   3396: 'Carrier 53 CB02122 Tripped', class No Acknowledgement, trigger "DB302_HMI_Faults_Carrier53_Faults_0" bit 3
   3397: 'Carrier 53 CB02123 Tripped', class No Acknowledgement, trigger "DB302_HMI_Faults_Carrier53_Faults_0" bit 4
   3398: 'Carrier 53 AUX1 CB Tripped', class No Acknowledgement, trigger "DB302_HMI_Faults_Carrier53_Faults_0" bit 5
   3399: 'Carrier 53 AUX2 CB Tripped', class No Acknowledgement, trigger "DB302_HMI_Faults_Carrier53_Faults_0" bit 6
   3400: 'Carrier 53 PLC Not Communicating', class No Acknowledgement, trigger "DB302_HMI_Faults_Carrier53_Faults_0" bit 7
   3401: 'Carrier 53 Safe Input Card Fault', class No Acknowledgement, trigger "DB302_HMI_Faults_Carrier53_Faults_0" bit 8
   3402: 'Carrier 53 Safe Output Card Fault', class No Acknowledgement, trigger "DB302_HMI_Faults_Carrier53_Faults_0" bit 9
   3403: 'Carrier 53 Standard Input Card Fault', class No Acknowledgement, trigger "DB302_HMI_Faults_Carrier53_Faults_0" bit 10
   3404: 'Carrier 53 Standard Output Card Fault', class No Acknowledgement, trigger "DB302_HMI_Faults_Carrier53_Faults_0" bit 11
   3405: 'Carrier 53 Encoder Position Fault', class No Acknowledgement, trigger "DB302_HMI_Faults_Carrier53_Faults_0" bit 12
   3406: 'Carrier 53 Encoder Internal Error', class No Acknowledgement, trigger "DB302_HMI_Faults_Carrier53_Faults_0" bit 13
   3407: 'Carrier 53 Encoder Comm Fault', class No Acknowledgement, trigger "DB302_HMI_Faults_Carrier53_Faults_0" bit 14
   3408: 'Carrier 53 HMI Comm Fault', class No Acknowledgement, trigger "DB302_HMI_Faults_Carrier53_Faults_0" bit 15
   3409: 'Carrier 53 Crash Detection Fault', class No Acknowledgement, trigger "DB302_HMI_Faults_Carrier53_Faults_1" bit 0
   3410: 'Carrier 53 Carrier Number Invalid', class No Acknowledgement, trigger "DB302_HMI_Faults_Carrier53_Faults_1" bit 1
   3411: 'Carrier 53 Drive: PROFINET configuration error', class No Acknowledgement, trigger "DB302_HMI_Faults_Carrier53_Faults_1" bit 2
   3412: 'Carrier 53 Drive: Error internal communications', class No Acknowledgement, trigger "DB302_HMI_Faults_Carrier53_Faults_1" bit 3
   3413: 'Carrier 53 Drive: Motor overtemperature', class No Acknowledgement, trigger "DB302_HMI_Faults_Carrier53_Faults_1" bit 4
   3414: 'Carrier 53 Drive: Motor overcurrent', class No Acknowledgement, trigger "DB302_HMI_Faults_Carrier53_Faults_1" bit 5
   3415: 'Carrier 53 Drive: Infeed or power unit not ready', class No Acknowledgement, trigger "DB302_HMI_Faults_Carrier53_Faults_1" bit 6
   3416: 'Carrier 53 Drive: Short-circuit/ground fault detected', class No Acknowledgement, trigger "DB302_HMI_Faults_Carrier53_Faults_1" bit 7
   3417: 'Carrier 53 Drive: PROFINET Setpoint timeout', class No Acknowledgement, trigger "DB302_HMI_Faults_Carrier53_Faults_1" bit 8
   3418: 'Carrier 53 Power unit: Overcurrent', class No Acknowledgement, trigger "DB302_HMI_Faults_Carrier53_Faults_1" bit 9
   3419: 'Carrier 53 Power unit: DC link voltage overvoltage', class No Acknowledgement, trigger "DB302_HMI_Faults_Carrier53_Faults_1" bit 10
   3420: 'Carrier 53 Power unit: DC link voltage undervoltage', class No Acknowledgement, trigger "DB302_HMI_Faults_Carrier53_Faults_1" bit 11
   3421: 'Carrier 53 Power unit: Line phase failure in main circuit', class No Acknowledgement, trigger "DB302_HMI_Faults_Carrier53_Faults_1" bit 12
   3422: 'Carrier 53 Power unit: Phase failure motor cable', class No Acknowledgement, trigger "DB302_HMI_Faults_Carrier53_Faults_1" bit 13
   3423: 'Carrier 53 Power unit: Ground fault', class No Acknowledgement, trigger "DB302_HMI_Faults_Carrier53_Faults_1" bit 14
   3424: 'Spare_Fault_3424', class No Acknowledgement, trigger "DB302_HMI_Faults_Carrier53_Faults_1" bit 15
   3425: 'Carrier 53 Motion Off Fault', class No Acknowledgement, trigger "DB302_HMI_Faults_Carrier53_Faults_2" bit 0
   3426: 'Carrier 53 Motion On Fault', class No Acknowledgement, trigger "DB302_HMI_Faults_Carrier53_Faults_2" bit 1
   3427: 'Carrier 53 Spacing Fault', class No Acknowledgement, trigger "DB302_HMI_Faults_Carrier53_Faults_2" bit 2
   3428: 'Carrier 53 Duplicate Carrier Number Fault', class No Acknowledgement, trigger "DB302_HMI_Faults_Carrier53_Faults_2" bit 3
   3429: 'Spare_Fault_3429', class No Acknowledgement, trigger "DB302_HMI_Faults_Carrier53_Faults_2" bit 4
   3430: 'Spare_Fault_3430', class No Acknowledgement, trigger "DB302_HMI_Faults_Carrier53_Faults_2" bit 5
   3431: 'Spare_Fault_3431', class No Acknowledgement, trigger "DB302_HMI_Faults_Carrier53_Faults_2" bit 6
   3432: 'Spare_Fault_3432', class No Acknowledgement, trigger "DB302_HMI_Faults_Carrier53_Faults_2" bit 7
   3433: 'Spare_Fault_3433', class No Acknowledgement, trigger "DB302_HMI_Faults_Carrier53_Faults_2" bit 8
   3434: 'Spare_Fault_3434', class No Acknowledgement, trigger "DB302_HMI_Faults_Carrier53_Faults_2" bit 9
   3435: 'Spare_Fault_3435', class No Acknowledgement, trigger "DB302_HMI_Faults_Carrier53_Faults_2" bit 10
   3436: 'Spare_Fault_3436', class No Acknowledgement, trigger "DB302_HMI_Faults_Carrier53_Faults_2" bit 11
   3437: 'Spare_Fault_3437', class No Acknowledgement, trigger "DB302_HMI_Faults_Carrier53_Faults_2" bit 12
   3438: 'Spare_Fault_3438', class No Acknowledgement, trigger "DB302_HMI_Faults_Carrier53_Faults_2" bit 13
   3439: 'Spare_Fault_3439', class No Acknowledgement, trigger "DB302_HMI_Faults_Carrier53_Faults_2" bit 14
   3440: 'Spare_Fault_3440', class No Acknowledgement, trigger "DB302_HMI_Faults_Carrier53_Faults_2" bit 15
   3441: 'Spare_Fault_3441', class No Acknowledgement, trigger "DB302_HMI_Faults_Carrier53_Faults_3" bit 0
   3442: 'Spare_Fault_3442', class No Acknowledgement, trigger "DB302_HMI_Faults_Carrier53_Faults_3" bit 1
   3443: 'Spare_Fault_3443', class No Acknowledgement, trigger "DB302_HMI_Faults_Carrier53_Faults_3" bit 2
   3444: 'Spare_Fault_3444', class No Acknowledgement, trigger "DB302_HMI_Faults_Carrier53_Faults_3" bit 3
   3445: 'Spare_Fault_3445', class No Acknowledgement, trigger "DB302_HMI_Faults_Carrier53_Faults_3" bit 4
   3446: 'Spare_Fault_3446', class No Acknowledgement, trigger "DB302_HMI_Faults_Carrier53_Faults_3" bit 5
   3447: 'Spare_Fault_3447', class No Acknowledgement, trigger "DB302_HMI_Faults_Carrier53_Faults_3" bit 6
   3448: 'Spare_Fault_3448', class No Acknowledgement, trigger "DB302_HMI_Faults_Carrier53_Faults_3" bit 7
   3449: 'Spare_Fault_3449', class No Acknowledgement, trigger "DB302_HMI_Faults_Carrier53_Faults_3" bit 8
   3450: 'Spare_Fault_3450', class No Acknowledgement, trigger "DB302_HMI_Faults_Carrier53_Faults_3" bit 9
   3451: 'Spare_Fault_3451', class No Acknowledgement, trigger "DB302_HMI_Faults_Carrier53_Faults_3" bit 10
   3452: 'Spare_Fault_3452', class No Acknowledgement, trigger "DB302_HMI_Faults_Carrier53_Faults_3" bit 11
   3453: 'Spare_Fault_3453', class No Acknowledgement, trigger "DB302_HMI_Faults_Carrier53_Faults_3" bit 12
   3454: 'Spare_Fault_3454', class No Acknowledgement, trigger "DB302_HMI_Faults_Carrier53_Faults_3" bit 13
   3455: 'Spare_Fault_3455', class No Acknowledgement, trigger "DB302_HMI_Faults_Carrier53_Faults_3" bit 14
   3456: 'Spare_Fault_3456', class No Acknowledgement, trigger "DB302_HMI_Faults_Carrier53_Faults_3" bit 15
   3457: 'Carrier 54 Disconnect Open Power Fault DI11.0', class No Acknowledgement, trigger "DB302_HMI_Faults_Carrier54_Faults_0" bit 0
   3458: 'Carrier 54 Drive Profinet Comm Fault', class No Acknowledgement, trigger "DB302_HMI_Faults_Carrier54_Faults_0" bit 1
   3459: 'Carrier 54 Production Stop Not Reset', class No Acknowledgement, trigger "DB302_HMI_Faults_Carrier54_Faults_0" bit 2
   3460: 'Carrier 54 CB02122 Tripped', class No Acknowledgement, trigger "DB302_HMI_Faults_Carrier54_Faults_0" bit 3
   3461: 'Carrier 54 CB02123 Tripped', class No Acknowledgement, trigger "DB302_HMI_Faults_Carrier54_Faults_0" bit 4
   3462: 'Carrier 54 AUX1 CB Tripped', class No Acknowledgement, trigger "DB302_HMI_Faults_Carrier54_Faults_0" bit 5
   3463: 'Carrier 54 AUX2 CB Tripped', class No Acknowledgement, trigger "DB302_HMI_Faults_Carrier54_Faults_0" bit 6
   3464: 'Carrier 54 PLC Not Communicating', class No Acknowledgement, trigger "DB302_HMI_Faults_Carrier54_Faults_0" bit 7
   3465: 'Carrier 54 Safe Input Card Fault', class No Acknowledgement, trigger "DB302_HMI_Faults_Carrier54_Faults_0" bit 8
   3466: 'Carrier 54 Safe Output Card Fault', class No Acknowledgement, trigger "DB302_HMI_Faults_Carrier54_Faults_0" bit 9
   3467: 'Carrier 54 Standard Input Card Fault', class No Acknowledgement, trigger "DB302_HMI_Faults_Carrier54_Faults_0" bit 10
   3468: 'Carrier 54 Standard Output Card Fault', class No Acknowledgement, trigger "DB302_HMI_Faults_Carrier54_Faults_0" bit 11
   3469: 'Carrier 54 Encoder Position Fault', class No Acknowledgement, trigger "DB302_HMI_Faults_Carrier54_Faults_0" bit 12
   3470: 'Carrier 54 Encoder Internal Error', class No Acknowledgement, trigger "DB302_HMI_Faults_Carrier54_Faults_0" bit 13
   3471: 'Carrier 54 Encoder Comm Fault', class No Acknowledgement, trigger "DB302_HMI_Faults_Carrier54_Faults_0" bit 14
   3472: 'Carrier 54 HMI Comm Fault', class No Acknowledgement, trigger "DB302_HMI_Faults_Carrier54_Faults_0" bit 15
   3473: 'Carrier 54 Crash Detection Fault', class No Acknowledgement, trigger "DB302_HMI_Faults_Carrier54_Faults_1" bit 0
   3474: 'Carrier 54 Carrier Number Invalid', class No Acknowledgement, trigger "DB302_HMI_Faults_Carrier54_Faults_1" bit 1
   3475: 'Carrier 54 Drive: PROFINET configuration error', class No Acknowledgement, trigger "DB302_HMI_Faults_Carrier54_Faults_1" bit 2
   3476: 'Carrier 54 Drive: Error internal communications', class No Acknowledgement, trigger "DB302_HMI_Faults_Carrier54_Faults_1" bit 3
   3477: 'Carrier 54 Drive: Motor overtemperature', class No Acknowledgement, trigger "DB302_HMI_Faults_Carrier54_Faults_1" bit 4
   3478: 'Carrier 54 Drive: Motor overcurrent', class No Acknowledgement, trigger "DB302_HMI_Faults_Carrier54_Faults_1" bit 5
   3479: 'Carrier 54 Drive: Infeed or power unit not ready', class No Acknowledgement, trigger "DB302_HMI_Faults_Carrier54_Faults_1" bit 6
   3480: 'Carrier 54 Drive: Short-circuit/ground fault detected', class No Acknowledgement, trigger "DB302_HMI_Faults_Carrier54_Faults_1" bit 7
   3481: 'Carrier 54 Drive: PROFINET Setpoint timeout', class No Acknowledgement, trigger "DB302_HMI_Faults_Carrier54_Faults_1" bit 8
   3482: 'Carrier 54 Power unit: Overcurrent', class No Acknowledgement, trigger "DB302_HMI_Faults_Carrier54_Faults_1" bit 9
   3483: 'Carrier 54 Power unit: DC link voltage overvoltage', class No Acknowledgement, trigger "DB302_HMI_Faults_Carrier54_Faults_1" bit 10
   3484: 'Carrier 54 Power unit: DC link voltage undervoltage', class No Acknowledgement, trigger "DB302_HMI_Faults_Carrier54_Faults_1" bit 11
   3485: 'Carrier 54 Power unit: Line phase failure in main circuit', class No Acknowledgement, trigger "DB302_HMI_Faults_Carrier54_Faults_1" bit 12
   3486: 'Carrier 54 Power unit: Phase failure motor cable', class No Acknowledgement, trigger "DB302_HMI_Faults_Carrier54_Faults_1" bit 13
   3487: 'Carrier 54 Power unit: Ground fault', class No Acknowledgement, trigger "DB302_HMI_Faults_Carrier54_Faults_1" bit 14
   3488: 'Spare_Fault_3488', class No Acknowledgement, trigger "DB302_HMI_Faults_Carrier54_Faults_1" bit 15
   3489: 'Carrier 54 Motion Off Fault', class No Acknowledgement, trigger "DB302_HMI_Faults_Carrier54_Faults_2" bit 0
   3490: 'Carrier 54 Motion On Fault', class No Acknowledgement, trigger "DB302_HMI_Faults_Carrier54_Faults_2" bit 1
   3491: 'Carrier 54 Spacing Fault', class No Acknowledgement, trigger "DB302_HMI_Faults_Carrier54_Faults_2" bit 2
   3492: 'Carrier 54 Duplicate Carrier Number Fault', class No Acknowledgement, trigger "DB302_HMI_Faults_Carrier54_Faults_2" bit 3
   3493: 'Spare_Fault_3493', class No Acknowledgement, trigger "DB302_HMI_Faults_Carrier54_Faults_2" bit 4
   3494: 'Spare_Fault_3494', class No Acknowledgement, trigger "DB302_HMI_Faults_Carrier54_Faults_2" bit 5
   3495: 'Spare_Fault_3495', class No Acknowledgement, trigger "DB302_HMI_Faults_Carrier54_Faults_2" bit 6
   3496: 'Spare_Fault_3496', class No Acknowledgement, trigger "DB302_HMI_Faults_Carrier54_Faults_2" bit 7
   3497: 'Spare_Fault_3497', class No Acknowledgement, trigger "DB302_HMI_Faults_Carrier54_Faults_2" bit 8
   3498: 'Spare_Fault_3498', class No Acknowledgement, trigger "DB302_HMI_Faults_Carrier54_Faults_2" bit 9
   3499: 'Spare_Fault_3499', class No Acknowledgement, trigger "DB302_HMI_Faults_Carrier54_Faults_2" bit 10
   3500: 'Spare_Fault_3500', class No Acknowledgement, trigger "DB302_HMI_Faults_Carrier54_Faults_2" bit 11
   3501: 'Spare_Fault_3501', class No Acknowledgement, trigger "DB302_HMI_Faults_Carrier54_Faults_2" bit 12
   3502: 'Spare_Fault_3502', class No Acknowledgement, trigger "DB302_HMI_Faults_Carrier54_Faults_2" bit 13
   3503: 'Spare_Fault_3503', class No Acknowledgement, trigger "DB302_HMI_Faults_Carrier54_Faults_2" bit 14
   3504: 'Spare_Fault_3504', class No Acknowledgement, trigger "DB302_HMI_Faults_Carrier54_Faults_2" bit 15
   3505: 'Spare_Fault_3505', class No Acknowledgement, trigger "DB302_HMI_Faults_Carrier54_Faults_3" bit 0
   3506: 'Spare_Fault_3506', class No Acknowledgement, trigger "DB302_HMI_Faults_Carrier54_Faults_3" bit 1
   3507: 'Spare_Fault_3507', class No Acknowledgement, trigger "DB302_HMI_Faults_Carrier54_Faults_3" bit 2
   3508: 'Spare_Fault_3508', class No Acknowledgement, trigger "DB302_HMI_Faults_Carrier54_Faults_3" bit 3
   3509: 'Spare_Fault_3509', class No Acknowledgement, trigger "DB302_HMI_Faults_Carrier54_Faults_3" bit 4
   3510: 'Spare_Fault_3510', class No Acknowledgement, trigger "DB302_HMI_Faults_Carrier54_Faults_3" bit 5
   3511: 'Spare_Fault_3511', class No Acknowledgement, trigger "DB302_HMI_Faults_Carrier54_Faults_3" bit 6
   3512: 'Spare_Fault_3512', class No Acknowledgement, trigger "DB302_HMI_Faults_Carrier54_Faults_3" bit 7
   3513: 'Spare_Fault_3513', class No Acknowledgement, trigger "DB302_HMI_Faults_Carrier54_Faults_3" bit 8
   3514: 'Spare_Fault_3514', class No Acknowledgement, trigger "DB302_HMI_Faults_Carrier54_Faults_3" bit 9
   3515: 'Spare_Fault_3515', class No Acknowledgement, trigger "DB302_HMI_Faults_Carrier54_Faults_3" bit 10
   3516: 'Spare_Fault_3516', class No Acknowledgement, trigger "DB302_HMI_Faults_Carrier54_Faults_3" bit 11
   3517: 'Spare_Fault_3517', class No Acknowledgement, trigger "DB302_HMI_Faults_Carrier54_Faults_3" bit 12
   3518: 'Spare_Fault_3518', class No Acknowledgement, trigger "DB302_HMI_Faults_Carrier54_Faults_3" bit 13
   3519: 'Spare_Fault_3519', class No Acknowledgement, trigger "DB302_HMI_Faults_Carrier54_Faults_3" bit 14
   3520: 'Spare_Fault_3520', class No Acknowledgement, trigger "DB302_HMI_Faults_Carrier54_Faults_3" bit 15
   3521: 'Carrier 55 Disconnect Open Power Fault DI11.0', class No Acknowledgement, trigger "DB302_HMI_Faults_Carrier55_Faults_0" bit 0
   3522: 'Carrier 55 Drive Profinet Comm Fault', class No Acknowledgement, trigger "DB302_HMI_Faults_Carrier55_Faults_0" bit 1
   3523: 'Carrier 55 Production Stop Not Reset', class No Acknowledgement, trigger "DB302_HMI_Faults_Carrier55_Faults_0" bit 2
   3524: 'Carrier 55 CB02122 Tripped', class No Acknowledgement, trigger "DB302_HMI_Faults_Carrier55_Faults_0" bit 3
   3525: 'Carrier 55 CB02123 Tripped', class No Acknowledgement, trigger "DB302_HMI_Faults_Carrier55_Faults_0" bit 4
   3526: 'Carrier 55 AUX1 CB Tripped', class No Acknowledgement, trigger "DB302_HMI_Faults_Carrier55_Faults_0" bit 5
   3527: 'Carrier 55 AUX2 CB Tripped', class No Acknowledgement, trigger "DB302_HMI_Faults_Carrier55_Faults_0" bit 6
   3528: 'Carrier 55 PLC Not Communicating', class No Acknowledgement, trigger "DB302_HMI_Faults_Carrier55_Faults_0" bit 7
   3529: 'Carrier 55 Safe Input Card Fault', class No Acknowledgement, trigger "DB302_HMI_Faults_Carrier55_Faults_0" bit 8
   3530: 'Carrier 55 Safe Output Card Fault', class No Acknowledgement, trigger "DB302_HMI_Faults_Carrier55_Faults_0" bit 9
   3531: 'Carrier 55 Standard Input Card Fault', class No Acknowledgement, trigger "DB302_HMI_Faults_Carrier55_Faults_0" bit 10
   3532: 'Carrier 55 Standard Output Card Fault', class No Acknowledgement, trigger "DB302_HMI_Faults_Carrier55_Faults_0" bit 11
   3533: 'Carrier 55 Encoder Position Fault', class No Acknowledgement, trigger "DB302_HMI_Faults_Carrier55_Faults_0" bit 12
   3534: 'Carrier 55 Encoder Internal Error', class No Acknowledgement, trigger "DB302_HMI_Faults_Carrier55_Faults_0" bit 13
   3535: 'Carrier 55 Encoder Comm Fault', class No Acknowledgement, trigger "DB302_HMI_Faults_Carrier55_Faults_0" bit 14
   3536: 'Carrier 55 HMI Comm Fault', class No Acknowledgement, trigger "DB302_HMI_Faults_Carrier55_Faults_0" bit 15
   3537: 'Carrier 55 Crash Detection Fault', class No Acknowledgement, trigger "DB302_HMI_Faults_Carrier55_Faults_1" bit 0
   3538: 'Carrier 55 Carrier Number Invalid', class No Acknowledgement, trigger "DB302_HMI_Faults_Carrier55_Faults_1" bit 1
   3539: 'Carrier 55 Drive: PROFINET configuration error', class No Acknowledgement, trigger "DB302_HMI_Faults_Carrier55_Faults_1" bit 2
   3540: 'Carrier 55 Drive: Error internal communications', class No Acknowledgement, trigger "DB302_HMI_Faults_Carrier55_Faults_1" bit 3
   3541: 'Carrier 55 Drive: Motor overtemperature', class No Acknowledgement, trigger "DB302_HMI_Faults_Carrier55_Faults_1" bit 4
   3542: 'Carrier 55 Drive: Motor overcurrent', class No Acknowledgement, trigger "DB302_HMI_Faults_Carrier55_Faults_1" bit 5
   3543: 'Carrier 55 Drive: Infeed or power unit not ready', class No Acknowledgement, trigger "DB302_HMI_Faults_Carrier55_Faults_1" bit 6
   3544: 'Carrier 55 Drive: Short-circuit/ground fault detected', class No Acknowledgement, trigger "DB302_HMI_Faults_Carrier55_Faults_1" bit 7
   3545: 'Carrier 55 Drive: PROFINET Setpoint timeout', class No Acknowledgement, trigger "DB302_HMI_Faults_Carrier55_Faults_1" bit 8
   3546: 'Carrier 55 Power unit: Overcurrent', class No Acknowledgement, trigger "DB302_HMI_Faults_Carrier55_Faults_1" bit 9
   3547: 'Carrier 55 Power unit: DC link voltage overvoltage', class No Acknowledgement, trigger "DB302_HMI_Faults_Carrier55_Faults_1" bit 10
   3548: 'Carrier 55 Power unit: DC link voltage undervoltage', class No Acknowledgement, trigger "DB302_HMI_Faults_Carrier55_Faults_1" bit 11
   3549: 'Carrier 55 Power unit: Line phase failure in main circuit', class No Acknowledgement, trigger "DB302_HMI_Faults_Carrier55_Faults_1" bit 12
   3550: 'Carrier 55 Power unit: Phase failure motor cable', class No Acknowledgement, trigger "DB302_HMI_Faults_Carrier55_Faults_1" bit 13
   3551: 'Carrier 55 Power unit: Ground fault', class No Acknowledgement, trigger "DB302_HMI_Faults_Carrier55_Faults_1" bit 14
   3552: 'Spare_Fault_3552', class No Acknowledgement, trigger "DB302_HMI_Faults_Carrier55_Faults_1" bit 15
   3553: 'Carrier 55 Motion Off Fault', class No Acknowledgement, trigger "DB302_HMI_Faults_Carrier55_Faults_2" bit 0
   3554: 'Carrier 55 Motion On Fault', class No Acknowledgement, trigger "DB302_HMI_Faults_Carrier55_Faults_2" bit 1
   3555: 'Carrier 55 Spacing Fault', class No Acknowledgement, trigger "DB302_HMI_Faults_Carrier55_Faults_2" bit 2
   3556: 'Carrier 55 Duplicate Carrier Number Fault', class No Acknowledgement, trigger "DB302_HMI_Faults_Carrier55_Faults_2" bit 3
   3557: 'Spare_Fault_3557', class No Acknowledgement, trigger "DB302_HMI_Faults_Carrier55_Faults_2" bit 4
   3558: 'Spare_Fault_3558', class No Acknowledgement, trigger "DB302_HMI_Faults_Carrier55_Faults_2" bit 5
   3559: 'Spare_Fault_3559', class No Acknowledgement, trigger "DB302_HMI_Faults_Carrier55_Faults_2" bit 6
   3560: 'Spare_Fault_3560', class No Acknowledgement, trigger "DB302_HMI_Faults_Carrier55_Faults_2" bit 7
   3561: 'Spare_Fault_3561', class No Acknowledgement, trigger "DB302_HMI_Faults_Carrier55_Faults_2" bit 8
   3562: 'Spare_Fault_3562', class No Acknowledgement, trigger "DB302_HMI_Faults_Carrier55_Faults_2" bit 9
   3563: 'Spare_Fault_3563', class No Acknowledgement, trigger "DB302_HMI_Faults_Carrier55_Faults_2" bit 10
   3564: 'Spare_Fault_3564', class No Acknowledgement, trigger "DB302_HMI_Faults_Carrier55_Faults_2" bit 11
   3565: 'Spare_Fault_3565', class No Acknowledgement, trigger "DB302_HMI_Faults_Carrier55_Faults_2" bit 12
   3566: 'Spare_Fault_3566', class No Acknowledgement, trigger "DB302_HMI_Faults_Carrier55_Faults_2" bit 13
   3567: 'Spare_Fault_3567', class No Acknowledgement, trigger "DB302_HMI_Faults_Carrier55_Faults_2" bit 14
   3568: 'Spare_Fault_3568', class No Acknowledgement, trigger "DB302_HMI_Faults_Carrier55_Faults_2" bit 15
   3569: 'Spare_Fault_3569', class No Acknowledgement, trigger "DB302_HMI_Faults_Carrier55_Faults_3" bit 0
   3570: 'Spare_Fault_3570', class No Acknowledgement, trigger "DB302_HMI_Faults_Carrier55_Faults_3" bit 1
   3571: 'Spare_Fault_3571', class No Acknowledgement, trigger "DB302_HMI_Faults_Carrier55_Faults_3" bit 2
   3572: 'Spare_Fault_3572', class No Acknowledgement, trigger "DB302_HMI_Faults_Carrier55_Faults_3" bit 3
   3573: 'Spare_Fault_3573', class No Acknowledgement, trigger "DB302_HMI_Faults_Carrier55_Faults_3" bit 4
   3574: 'Spare_Fault_3574', class No Acknowledgement, trigger "DB302_HMI_Faults_Carrier55_Faults_3" bit 5
   3575: 'Spare_Fault_3575', class No Acknowledgement, trigger "DB302_HMI_Faults_Carrier55_Faults_3" bit 6
   3576: 'Spare_Fault_3576', class No Acknowledgement, trigger "DB302_HMI_Faults_Carrier55_Faults_3" bit 7
   3577: 'Spare_Fault_3577', class No Acknowledgement, trigger "DB302_HMI_Faults_Carrier55_Faults_3" bit 8
   3578: 'Spare_Fault_3578', class No Acknowledgement, trigger "DB302_HMI_Faults_Carrier55_Faults_3" bit 9
   3579: 'Spare_Fault_3579', class No Acknowledgement, trigger "DB302_HMI_Faults_Carrier55_Faults_3" bit 10
   3580: 'Spare_Fault_3580', class No Acknowledgement, trigger "DB302_HMI_Faults_Carrier55_Faults_3" bit 11
   3581: 'Spare_Fault_3581', class No Acknowledgement, trigger "DB302_HMI_Faults_Carrier55_Faults_3" bit 12
   3582: 'Spare_Fault_3582', class No Acknowledgement, trigger "DB302_HMI_Faults_Carrier55_Faults_3" bit 13
   3583: 'Spare_Fault_3583', class No Acknowledgement, trigger "DB302_HMI_Faults_Carrier55_Faults_3" bit 14
   3584: 'Spare_Fault_3584', class No Acknowledgement, trigger "DB302_HMI_Faults_Carrier55_Faults_3" bit 15
   3585: 'Carrier 56 Disconnect Open Power Fault DI11.0', class No Acknowledgement, trigger "DB302_HMI_Faults_Carrier56_Faults_0" bit 0
   3586: 'Carrier 56 Drive Profinet Comm Fault', class No Acknowledgement, trigger "DB302_HMI_Faults_Carrier56_Faults_0" bit 1
   3587: 'Carrier 56 Production Stop Not Reset', class No Acknowledgement, trigger "DB302_HMI_Faults_Carrier56_Faults_0" bit 2
   3588: 'Carrier 56 CB02122 Tripped', class No Acknowledgement, trigger "DB302_HMI_Faults_Carrier56_Faults_0" bit 3
   3589: 'Carrier 56 CB02123 Tripped', class No Acknowledgement, trigger "DB302_HMI_Faults_Carrier56_Faults_0" bit 4
   3590: 'Carrier 56 AUX1 CB Tripped', class No Acknowledgement, trigger "DB302_HMI_Faults_Carrier56_Faults_0" bit 5
   3591: 'Carrier 56 AUX2 CB Tripped', class No Acknowledgement, trigger "DB302_HMI_Faults_Carrier56_Faults_0" bit 6
   3592: 'Carrier 56 PLC Not Communicating', class No Acknowledgement, trigger "DB302_HMI_Faults_Carrier56_Faults_0" bit 7
   3593: 'Carrier 56 Safe Input Card Fault', class No Acknowledgement, trigger "DB302_HMI_Faults_Carrier56_Faults_0" bit 8
   3594: 'Carrier 56 Safe Output Card Fault', class No Acknowledgement, trigger "DB302_HMI_Faults_Carrier56_Faults_0" bit 9
   3595: 'Carrier 56 Standard Input Card Fault', class No Acknowledgement, trigger "DB302_HMI_Faults_Carrier56_Faults_0" bit 10
   3596: 'Carrier 56 Standard Output Card Fault', class No Acknowledgement, trigger "DB302_HMI_Faults_Carrier56_Faults_0" bit 11
   3597: 'Carrier 56 Encoder Position Fault', class No Acknowledgement, trigger "DB302_HMI_Faults_Carrier56_Faults_0" bit 12
   3598: 'Carrier 56 Encoder Internal Error', class No Acknowledgement, trigger "DB302_HMI_Faults_Carrier56_Faults_0" bit 13
   3599: 'Carrier 56 Encoder Comm Fault', class No Acknowledgement, trigger "DB302_HMI_Faults_Carrier56_Faults_0" bit 14
   3600: 'Carrier 56 HMI Comm Fault', class No Acknowledgement, trigger "DB302_HMI_Faults_Carrier56_Faults_0" bit 15
   3601: 'Carrier 56 Crash Detection Fault', class No Acknowledgement, trigger "DB302_HMI_Faults_Carrier56_Faults_1" bit 0
   3602: 'Carrier 56 Carrier Number Invalid', class No Acknowledgement, trigger "DB302_HMI_Faults_Carrier56_Faults_1" bit 1
   3603: 'Carrier 56 Drive: PROFINET configuration error', class No Acknowledgement, trigger "DB302_HMI_Faults_Carrier56_Faults_1" bit 2
   3604: 'Carrier 56 Drive: Error internal communications', class No Acknowledgement, trigger "DB302_HMI_Faults_Carrier56_Faults_1" bit 3
   3605: 'Carrier 56 Drive: Motor overtemperature', class No Acknowledgement, trigger "DB302_HMI_Faults_Carrier56_Faults_1" bit 4
   3606: 'Carrier 56 Drive: Motor overcurrent', class No Acknowledgement, trigger "DB302_HMI_Faults_Carrier56_Faults_1" bit 5
   3607: 'Carrier 56 Drive: Infeed or power unit not ready', class No Acknowledgement, trigger "DB302_HMI_Faults_Carrier56_Faults_1" bit 6
   3608: 'Carrier 56 Drive: Short-circuit/ground fault detected', class No Acknowledgement, trigger "DB302_HMI_Faults_Carrier56_Faults_1" bit 7
   3609: 'Carrier 56 Drive: PROFINET Setpoint timeout', class No Acknowledgement, trigger "DB302_HMI_Faults_Carrier56_Faults_1" bit 8
   3610: 'Carrier 56 Power unit: Overcurrent', class No Acknowledgement, trigger "DB302_HMI_Faults_Carrier56_Faults_1" bit 9
   3611: 'Carrier 56 Power unit: DC link voltage overvoltage', class No Acknowledgement, trigger "DB302_HMI_Faults_Carrier56_Faults_1" bit 10
   3612: 'Carrier 56 Power unit: DC link voltage undervoltage', class No Acknowledgement, trigger "DB302_HMI_Faults_Carrier56_Faults_1" bit 11
   3613: 'Carrier 56 Power unit: Line phase failure in main circuit', class No Acknowledgement, trigger "DB302_HMI_Faults_Carrier56_Faults_1" bit 12
   3614: 'Carrier 56 Power unit: Phase failure motor cable', class No Acknowledgement, trigger "DB302_HMI_Faults_Carrier56_Faults_1" bit 13
   3615: 'Carrier 56 Power unit: Ground fault', class No Acknowledgement, trigger "DB302_HMI_Faults_Carrier56_Faults_1" bit 14
   3616: 'Spare_Fault_3616', class No Acknowledgement, trigger "DB302_HMI_Faults_Carrier56_Faults_1" bit 15
   3617: 'Carrier 56 Motion Off Fault', class No Acknowledgement, trigger "DB302_HMI_Faults_Carrier56_Faults_2" bit 0
   3618: 'Carrier 56 Motion On Fault', class No Acknowledgement, trigger "DB302_HMI_Faults_Carrier56_Faults_2" bit 1
   3619: 'Carrier 56 Spacing Fault', class No Acknowledgement, trigger "DB302_HMI_Faults_Carrier56_Faults_2" bit 2
   3620: 'Carrier 56 Duplicate Carrier Number Fault', class No Acknowledgement, trigger "DB302_HMI_Faults_Carrier56_Faults_2" bit 3
   3621: 'Spare_Fault_3621', class No Acknowledgement, trigger "DB302_HMI_Faults_Carrier56_Faults_2" bit 4
   3622: 'Spare_Fault_3622', class No Acknowledgement, trigger "DB302_HMI_Faults_Carrier56_Faults_2" bit 5
   3623: 'Spare_Fault_3623', class No Acknowledgement, trigger "DB302_HMI_Faults_Carrier56_Faults_2" bit 6
   3624: 'Spare_Fault_3624', class No Acknowledgement, trigger "DB302_HMI_Faults_Carrier56_Faults_2" bit 7
   3625: 'Spare_Fault_3625', class No Acknowledgement, trigger "DB302_HMI_Faults_Carrier56_Faults_2" bit 8
   3626: 'Spare_Fault_3626', class No Acknowledgement, trigger "DB302_HMI_Faults_Carrier56_Faults_2" bit 9
   3627: 'Spare_Fault_3627', class No Acknowledgement, trigger "DB302_HMI_Faults_Carrier56_Faults_2" bit 10
   3628: 'Spare_Fault_3628', class No Acknowledgement, trigger "DB302_HMI_Faults_Carrier56_Faults_2" bit 11
   3629: 'Spare_Fault_3629', class No Acknowledgement, trigger "DB302_HMI_Faults_Carrier56_Faults_2" bit 12
   3630: 'Spare_Fault_3630', class No Acknowledgement, trigger "DB302_HMI_Faults_Carrier56_Faults_2" bit 13
   3631: 'Spare_Fault_3631', class No Acknowledgement, trigger "DB302_HMI_Faults_Carrier56_Faults_2" bit 14
   3632: 'Spare_Fault_3632', class No Acknowledgement, trigger "DB302_HMI_Faults_Carrier56_Faults_2" bit 15
   3633: 'Spare_Fault_3633', class No Acknowledgement, trigger "DB302_HMI_Faults_Carrier56_Faults_3" bit 0
   3634: 'Spare_Fault_3634', class No Acknowledgement, trigger "DB302_HMI_Faults_Carrier56_Faults_3" bit 1
   3635: 'Spare_Fault_3635', class No Acknowledgement, trigger "DB302_HMI_Faults_Carrier56_Faults_3" bit 2
   3636: 'Spare_Fault_3636', class No Acknowledgement, trigger "DB302_HMI_Faults_Carrier56_Faults_3" bit 3
   3637: 'Spare_Fault_3637', class No Acknowledgement, trigger "DB302_HMI_Faults_Carrier56_Faults_3" bit 4
   3638: 'Spare_Fault_3638', class No Acknowledgement, trigger "DB302_HMI_Faults_Carrier56_Faults_3" bit 5
   3639: 'Spare_Fault_3639', class No Acknowledgement, trigger "DB302_HMI_Faults_Carrier56_Faults_3" bit 6
   3640: 'Spare_Fault_3640', class No Acknowledgement, trigger "DB302_HMI_Faults_Carrier56_Faults_3" bit 7
   3641: 'Spare_Fault_3641', class No Acknowledgement, trigger "DB302_HMI_Faults_Carrier56_Faults_3" bit 8
   3642: 'Spare_Fault_3642', class No Acknowledgement, trigger "DB302_HMI_Faults_Carrier56_Faults_3" bit 9
   3643: 'Spare_Fault_3643', class No Acknowledgement, trigger "DB302_HMI_Faults_Carrier56_Faults_3" bit 10
   3644: 'Spare_Fault_3644', class No Acknowledgement, trigger "DB302_HMI_Faults_Carrier56_Faults_3" bit 11
   3645: 'Spare_Fault_3645', class No Acknowledgement, trigger "DB302_HMI_Faults_Carrier56_Faults_3" bit 12
   3646: 'Spare_Fault_3646', class No Acknowledgement, trigger "DB302_HMI_Faults_Carrier56_Faults_3" bit 13
   3647: 'Spare_Fault_3647', class No Acknowledgement, trigger "DB302_HMI_Faults_Carrier56_Faults_3" bit 14
   3648: 'Spare_Fault_3648', class No Acknowledgement, trigger "DB302_HMI_Faults_Carrier56_Faults_3" bit 15
   3649: 'Carrier 57 Disconnect Open Power Fault DI11.0', class No Acknowledgement, trigger "DB302_HMI_Faults_Carrier57_Faults_0" bit 0
   3650: 'Carrier 57 Drive Profinet Comm Fault', class No Acknowledgement, trigger "DB302_HMI_Faults_Carrier57_Faults_0" bit 1
   3651: 'Carrier 57 Production Stop Not Reset', class No Acknowledgement, trigger "DB302_HMI_Faults_Carrier57_Faults_0" bit 2
   3652: 'Carrier 57 CB02122 Tripped', class No Acknowledgement, trigger "DB302_HMI_Faults_Carrier57_Faults_0" bit 3
   3653: 'Carrier 57 CB02123 Tripped', class No Acknowledgement, trigger "DB302_HMI_Faults_Carrier57_Faults_0" bit 4
   3654: 'Carrier 57 AUX1 CB Tripped', class No Acknowledgement, trigger "DB302_HMI_Faults_Carrier57_Faults_0" bit 5
   3655: 'Carrier 57 AUX2 CB Tripped', class No Acknowledgement, trigger "DB302_HMI_Faults_Carrier57_Faults_0" bit 6
   3656: 'Carrier 57 PLC Not Communicating', class No Acknowledgement, trigger "DB302_HMI_Faults_Carrier57_Faults_0" bit 7
   3657: 'Carrier 57 Safe Input Card Fault', class No Acknowledgement, trigger "DB302_HMI_Faults_Carrier57_Faults_0" bit 8
   3658: 'Carrier 57 Safe Output Card Fault', class No Acknowledgement, trigger "DB302_HMI_Faults_Carrier57_Faults_0" bit 9
   3659: 'Carrier 57 Standard Input Card Fault', class No Acknowledgement, trigger "DB302_HMI_Faults_Carrier57_Faults_0" bit 10
   3660: 'Carrier 57 Standard Output Card Fault', class No Acknowledgement, trigger "DB302_HMI_Faults_Carrier57_Faults_0" bit 11
   3661: 'Carrier 57 Encoder Position Fault', class No Acknowledgement, trigger "DB302_HMI_Faults_Carrier57_Faults_0" bit 12
   3662: 'Carrier 57 Encoder Internal Error', class No Acknowledgement, trigger "DB302_HMI_Faults_Carrier57_Faults_0" bit 13
   3663: 'Carrier 57 Encoder Comm Fault', class No Acknowledgement, trigger "DB302_HMI_Faults_Carrier57_Faults_0" bit 14
   3664: 'Carrier 57 HMI Comm Fault', class No Acknowledgement, trigger "DB302_HMI_Faults_Carrier57_Faults_0" bit 15
   3665: 'Carrier 57 Crash Detection Fault', class No Acknowledgement, trigger "DB302_HMI_Faults_Carrier57_Faults_1" bit 0
   3666: 'Carrier 57 Carrier Number Invalid', class No Acknowledgement, trigger "DB302_HMI_Faults_Carrier57_Faults_1" bit 1
   3667: 'Carrier 57 Drive: PROFINET configuration error', class No Acknowledgement, trigger "DB302_HMI_Faults_Carrier57_Faults_1" bit 2
   3668: 'Carrier 57 Drive: Error internal communications', class No Acknowledgement, trigger "DB302_HMI_Faults_Carrier57_Faults_1" bit 3
   3669: 'Carrier 57 Drive: Motor overtemperature', class No Acknowledgement, trigger "DB302_HMI_Faults_Carrier57_Faults_1" bit 4
   3670: 'Carrier 57 Drive: Motor overcurrent', class No Acknowledgement, trigger "DB302_HMI_Faults_Carrier57_Faults_1" bit 5
   3671: 'Carrier 57 Drive: Infeed or power unit not ready', class No Acknowledgement, trigger "DB302_HMI_Faults_Carrier57_Faults_1" bit 6
   3672: 'Carrier 57 Drive: Short-circuit/ground fault detected', class No Acknowledgement, trigger "DB302_HMI_Faults_Carrier57_Faults_1" bit 7
   3673: 'Carrier 57 Drive: PROFINET Setpoint timeout', class No Acknowledgement, trigger "DB302_HMI_Faults_Carrier57_Faults_1" bit 8
   3674: 'Carrier 57 Power unit: Overcurrent', class No Acknowledgement, trigger "DB302_HMI_Faults_Carrier57_Faults_1" bit 9
   3675: 'Carrier 57 Power unit: DC link voltage overvoltage', class No Acknowledgement, trigger "DB302_HMI_Faults_Carrier57_Faults_1" bit 10
   3676: 'Carrier 57 Power unit: DC link voltage undervoltage', class No Acknowledgement, trigger "DB302_HMI_Faults_Carrier57_Faults_1" bit 11
   3677: 'Carrier 57 Power unit: Line phase failure in main circuit', class No Acknowledgement, trigger "DB302_HMI_Faults_Carrier57_Faults_1" bit 12
   3678: 'Carrier 57 Power unit: Phase failure motor cable', class No Acknowledgement, trigger "DB302_HMI_Faults_Carrier57_Faults_1" bit 13
   3679: 'Carrier 57 Power unit: Ground fault', class No Acknowledgement, trigger "DB302_HMI_Faults_Carrier57_Faults_1" bit 14
   3680: 'Spare_Fault_3680', class No Acknowledgement, trigger "DB302_HMI_Faults_Carrier57_Faults_1" bit 15
   3681: 'Carrier 57 Motion Off Fault', class No Acknowledgement, trigger "DB302_HMI_Faults_Carrier57_Faults_2" bit 0
   3682: 'Carrier 57 Motion On Fault', class No Acknowledgement, trigger "DB302_HMI_Faults_Carrier57_Faults_2" bit 1
   3683: 'Carrier 57 Spacing Fault', class No Acknowledgement, trigger "DB302_HMI_Faults_Carrier57_Faults_2" bit 2
   3684: 'Carrier 57 Duplicate Carrier Number Fault', class No Acknowledgement, trigger "DB302_HMI_Faults_Carrier57_Faults_2" bit 3
   3685: 'Spare_Fault_3685', class No Acknowledgement, trigger "DB302_HMI_Faults_Carrier57_Faults_2" bit 4
   3686: 'Spare_Fault_3686', class No Acknowledgement, trigger "DB302_HMI_Faults_Carrier57_Faults_2" bit 5
   3687: 'Spare_Fault_3687', class No Acknowledgement, trigger "DB302_HMI_Faults_Carrier57_Faults_2" bit 6
   3688: 'Spare_Fault_3688', class No Acknowledgement, trigger "DB302_HMI_Faults_Carrier57_Faults_2" bit 7
   3689: 'Spare_Fault_3689', class No Acknowledgement, trigger "DB302_HMI_Faults_Carrier57_Faults_2" bit 8
   3690: 'Spare_Fault_3690', class No Acknowledgement, trigger "DB302_HMI_Faults_Carrier57_Faults_2" bit 9
   3691: 'Spare_Fault_3691', class No Acknowledgement, trigger "DB302_HMI_Faults_Carrier57_Faults_2" bit 10
   3692: 'Spare_Fault_3692', class No Acknowledgement, trigger "DB302_HMI_Faults_Carrier57_Faults_2" bit 11
   3693: 'Spare_Fault_3693', class No Acknowledgement, trigger "DB302_HMI_Faults_Carrier57_Faults_2" bit 12
   3694: 'Spare_Fault_3694', class No Acknowledgement, trigger "DB302_HMI_Faults_Carrier57_Faults_2" bit 13
   3695: 'Spare_Fault_3695', class No Acknowledgement, trigger "DB302_HMI_Faults_Carrier57_Faults_2" bit 14
   3696: 'Spare_Fault_3696', class No Acknowledgement, trigger "DB302_HMI_Faults_Carrier57_Faults_2" bit 15
   3697: 'Spare_Fault_3697', class No Acknowledgement, trigger "DB302_HMI_Faults_Carrier57_Faults_3" bit 0
   3698: 'Spare_Fault_3698', class No Acknowledgement, trigger "DB302_HMI_Faults_Carrier57_Faults_3" bit 1
   3699: 'Spare_Fault_3699', class No Acknowledgement, trigger "DB302_HMI_Faults_Carrier57_Faults_3" bit 2
   3700: 'Spare_Fault_3700', class No Acknowledgement, trigger "DB302_HMI_Faults_Carrier57_Faults_3" bit 3
   3701: 'Spare_Fault_3701', class No Acknowledgement, trigger "DB302_HMI_Faults_Carrier57_Faults_3" bit 4
   3702: 'Spare_Fault_3702', class No Acknowledgement, trigger "DB302_HMI_Faults_Carrier57_Faults_3" bit 5
   3703: 'Spare_Fault_3703', class No Acknowledgement, trigger "DB302_HMI_Faults_Carrier57_Faults_3" bit 6
   3704: 'Spare_Fault_3704', class No Acknowledgement, trigger "DB302_HMI_Faults_Carrier57_Faults_3" bit 7
   3705: 'Spare_Fault_3705', class No Acknowledgement, trigger "DB302_HMI_Faults_Carrier57_Faults_3" bit 8
   3706: 'Spare_Fault_3706', class No Acknowledgement, trigger "DB302_HMI_Faults_Carrier57_Faults_3" bit 9
   3707: 'Spare_Fault_3707', class No Acknowledgement, trigger "DB302_HMI_Faults_Carrier57_Faults_3" bit 10
   3708: 'Spare_Fault_3708', class No Acknowledgement, trigger "DB302_HMI_Faults_Carrier57_Faults_3" bit 11
   3709: 'Spare_Fault_3709', class No Acknowledgement, trigger "DB302_HMI_Faults_Carrier57_Faults_3" bit 12
   3710: 'Spare_Fault_3710', class No Acknowledgement, trigger "DB302_HMI_Faults_Carrier57_Faults_3" bit 13
   3711: 'Spare_Fault_3711', class No Acknowledgement, trigger "DB302_HMI_Faults_Carrier57_Faults_3" bit 14
   3712: 'Spare_Fault_3712', class No Acknowledgement, trigger "DB302_HMI_Faults_Carrier57_Faults_3" bit 15
   3713: 'Carrier 58 Disconnect Open Power Fault DI11.0', class No Acknowledgement, trigger "DB302_HMI_Faults_Carrier58_Faults_0" bit 0
   3714: 'Carrier 58 Drive Profinet Comm Fault', class No Acknowledgement, trigger "DB302_HMI_Faults_Carrier58_Faults_0" bit 1
   3715: 'Carrier 58 Production Stop Not Reset', class No Acknowledgement, trigger "DB302_HMI_Faults_Carrier58_Faults_0" bit 2
   3716: 'Carrier 58 CB02122 Tripped', class No Acknowledgement, trigger "DB302_HMI_Faults_Carrier58_Faults_0" bit 3
   3717: 'Carrier 58 CB02123 Tripped', class No Acknowledgement, trigger "DB302_HMI_Faults_Carrier58_Faults_0" bit 4
   3718: 'Carrier 58 AUX1 CB Tripped', class No Acknowledgement, trigger "DB302_HMI_Faults_Carrier58_Faults_0" bit 5
   3719: 'Carrier 58 AUX2 CB Tripped', class No Acknowledgement, trigger "DB302_HMI_Faults_Carrier58_Faults_0" bit 6
   3720: 'Carrier 58 PLC Not Communicating', class No Acknowledgement, trigger "DB302_HMI_Faults_Carrier58_Faults_0" bit 7
   3721: 'Carrier 58 Safe Input Card Fault', class No Acknowledgement, trigger "DB302_HMI_Faults_Carrier58_Faults_0" bit 8
   3722: 'Carrier 58 Safe Output Card Fault', class No Acknowledgement, trigger "DB302_HMI_Faults_Carrier58_Faults_0" bit 9
   3723: 'Carrier 58 Standard Input Card Fault', class No Acknowledgement, trigger "DB302_HMI_Faults_Carrier58_Faults_0" bit 10
   3724: 'Carrier 58 Standard Output Card Fault', class No Acknowledgement, trigger "DB302_HMI_Faults_Carrier58_Faults_0" bit 11
   3725: 'Carrier 58 Encoder Position Fault', class No Acknowledgement, trigger "DB302_HMI_Faults_Carrier58_Faults_0" bit 12
   3726: 'Carrier 58 Encoder Internal Error', class No Acknowledgement, trigger "DB302_HMI_Faults_Carrier58_Faults_0" bit 13
   3727: 'Carrier 58 Encoder Comm Fault', class No Acknowledgement, trigger "DB302_HMI_Faults_Carrier58_Faults_0" bit 14
   3728: 'Carrier 58 HMI Comm Fault', class No Acknowledgement, trigger "DB302_HMI_Faults_Carrier58_Faults_0" bit 15
   3729: 'Carrier 58 Crash Detection Fault', class No Acknowledgement, trigger "DB302_HMI_Faults_Carrier58_Faults_1" bit 0
   3730: 'Carrier 58 Carrier Number Invalid', class No Acknowledgement, trigger "DB302_HMI_Faults_Carrier58_Faults_1" bit 1
   3731: 'Carrier 58 Drive: PROFINET configuration error', class No Acknowledgement, trigger "DB302_HMI_Faults_Carrier58_Faults_1" bit 2
   3732: 'Carrier 58 Drive: Error internal communications', class No Acknowledgement, trigger "DB302_HMI_Faults_Carrier58_Faults_1" bit 3
   3733: 'Carrier 58 Drive: Motor overtemperature', class No Acknowledgement, trigger "DB302_HMI_Faults_Carrier58_Faults_1" bit 4
   3734: 'Carrier 58 Drive: Motor overcurrent', class No Acknowledgement, trigger "DB302_HMI_Faults_Carrier58_Faults_1" bit 5
   3735: 'Carrier 58 Drive: Infeed or power unit not ready', class No Acknowledgement, trigger "DB302_HMI_Faults_Carrier58_Faults_1" bit 6
   3736: 'Carrier 58 Drive: Short-circuit/ground fault detected', class No Acknowledgement, trigger "DB302_HMI_Faults_Carrier58_Faults_1" bit 7
   3737: 'Carrier 58 Drive: PROFINET Setpoint timeout', class No Acknowledgement, trigger "DB302_HMI_Faults_Carrier58_Faults_1" bit 8
   3738: 'Carrier 58 Power unit: Overcurrent', class No Acknowledgement, trigger "DB302_HMI_Faults_Carrier58_Faults_1" bit 9
   3739: 'Carrier 58 Power unit: DC link voltage overvoltage', class No Acknowledgement, trigger "DB302_HMI_Faults_Carrier58_Faults_1" bit 10
   3740: 'Carrier 58 Power unit: DC link voltage undervoltage', class No Acknowledgement, trigger "DB302_HMI_Faults_Carrier58_Faults_1" bit 11
   3741: 'Carrier 58 Power unit: Line phase failure in main circuit', class No Acknowledgement, trigger "DB302_HMI_Faults_Carrier58_Faults_1" bit 12
   3742: 'Carrier 58 Power unit: Phase failure motor cable', class No Acknowledgement, trigger "DB302_HMI_Faults_Carrier58_Faults_1" bit 13
   3743: 'Carrier 58 Power unit: Ground fault', class No Acknowledgement, trigger "DB302_HMI_Faults_Carrier58_Faults_1" bit 14
   3744: 'Spare_Fault_3744', class No Acknowledgement, trigger "DB302_HMI_Faults_Carrier58_Faults_1" bit 15
   3745: 'Carrier 58 Motion Off Fault', class No Acknowledgement, trigger "DB302_HMI_Faults_Carrier58_Faults_2" bit 0
   3746: 'Carrier 58 Motion On Fault', class No Acknowledgement, trigger "DB302_HMI_Faults_Carrier58_Faults_2" bit 1
   3747: 'Carrier 58 Spacing Fault', class No Acknowledgement, trigger "DB302_HMI_Faults_Carrier58_Faults_2" bit 2
   3748: 'Carrier 58 Duplicate Carrier Number Fault', class No Acknowledgement, trigger "DB302_HMI_Faults_Carrier58_Faults_2" bit 3
   3749: 'Spare_Fault_3749', class No Acknowledgement, trigger "DB302_HMI_Faults_Carrier58_Faults_2" bit 4
   3750: 'Spare_Fault_3750', class No Acknowledgement, trigger "DB302_HMI_Faults_Carrier58_Faults_2" bit 5
   3751: 'Spare_Fault_3751', class No Acknowledgement, trigger "DB302_HMI_Faults_Carrier58_Faults_2" bit 6
   3752: 'Spare_Fault_3752', class No Acknowledgement, trigger "DB302_HMI_Faults_Carrier58_Faults_2" bit 7
   3753: 'Spare_Fault_3753', class No Acknowledgement, trigger "DB302_HMI_Faults_Carrier58_Faults_2" bit 8
   3754: 'Spare_Fault_3754', class No Acknowledgement, trigger "DB302_HMI_Faults_Carrier58_Faults_2" bit 9
   3755: 'Spare_Fault_3755', class No Acknowledgement, trigger "DB302_HMI_Faults_Carrier58_Faults_2" bit 10
   3756: 'Spare_Fault_3756', class No Acknowledgement, trigger "DB302_HMI_Faults_Carrier58_Faults_2" bit 11
   3757: 'Spare_Fault_3757', class No Acknowledgement, trigger "DB302_HMI_Faults_Carrier58_Faults_2" bit 12
   3758: 'Spare_Fault_3758', class No Acknowledgement, trigger "DB302_HMI_Faults_Carrier58_Faults_2" bit 13
   3759: 'Spare_Fault_3759', class No Acknowledgement, trigger "DB302_HMI_Faults_Carrier58_Faults_2" bit 14
   3760: 'Spare_Fault_3760', class No Acknowledgement, trigger "DB302_HMI_Faults_Carrier58_Faults_2" bit 15
   3761: 'Spare_Fault_3761', class No Acknowledgement, trigger "DB302_HMI_Faults_Carrier58_Faults_3" bit 0
   3762: 'Spare_Fault_3762', class No Acknowledgement, trigger "DB302_HMI_Faults_Carrier58_Faults_3" bit 1
   3763: 'Spare_Fault_3763', class No Acknowledgement, trigger "DB302_HMI_Faults_Carrier58_Faults_3" bit 2
   3764: 'Spare_Fault_3764', class No Acknowledgement, trigger "DB302_HMI_Faults_Carrier58_Faults_3" bit 3
   3765: 'Spare_Fault_3765', class No Acknowledgement, trigger "DB302_HMI_Faults_Carrier58_Faults_3" bit 4
   3766: 'Spare_Fault_3766', class No Acknowledgement, trigger "DB302_HMI_Faults_Carrier58_Faults_3" bit 5
   3767: 'Spare_Fault_3767', class No Acknowledgement, trigger "DB302_HMI_Faults_Carrier58_Faults_3" bit 6
   3768: 'Spare_Fault_3768', class No Acknowledgement, trigger "DB302_HMI_Faults_Carrier58_Faults_3" bit 7
   3769: 'Spare_Fault_3769', class No Acknowledgement, trigger "DB302_HMI_Faults_Carrier58_Faults_3" bit 8
   3770: 'Spare_Fault_3770', class No Acknowledgement, trigger "DB302_HMI_Faults_Carrier58_Faults_3" bit 9
   3771: 'Spare_Fault_3771', class No Acknowledgement, trigger "DB302_HMI_Faults_Carrier58_Faults_3" bit 10
   3772: 'Spare_Fault_3772', class No Acknowledgement, trigger "DB302_HMI_Faults_Carrier58_Faults_3" bit 11
   3773: 'Spare_Fault_3773', class No Acknowledgement, trigger "DB302_HMI_Faults_Carrier58_Faults_3" bit 12
   3774: 'Spare_Fault_3774', class No Acknowledgement, trigger "DB302_HMI_Faults_Carrier58_Faults_3" bit 13
   3775: 'Spare_Fault_3775', class No Acknowledgement, trigger "DB302_HMI_Faults_Carrier58_Faults_3" bit 14
   3776: 'Spare_Fault_3776', class No Acknowledgement, trigger "DB302_HMI_Faults_Carrier58_Faults_3" bit 15
   3777: 'Carrier 59 Disconnect Open Power Fault DI11.0', class No Acknowledgement, trigger "DB302_HMI_Faults_Carrier59_Faults_0" bit 0
   3778: 'Carrier 59 Drive Profinet Comm Fault', class No Acknowledgement, trigger "DB302_HMI_Faults_Carrier59_Faults_0" bit 1
   3779: 'Carrier 59 Production Stop Not Reset', class No Acknowledgement, trigger "DB302_HMI_Faults_Carrier59_Faults_0" bit 2
   3780: 'Carrier 59 CB02122 Tripped', class No Acknowledgement, trigger "DB302_HMI_Faults_Carrier59_Faults_0" bit 3
   3781: 'Carrier 59 CB02123 Tripped', class No Acknowledgement, trigger "DB302_HMI_Faults_Carrier59_Faults_0" bit 4
   3782: 'Carrier 59 AUX1 CB Tripped', class No Acknowledgement, trigger "DB302_HMI_Faults_Carrier59_Faults_0" bit 5
   3783: 'Carrier 59 AUX2 CB Tripped', class No Acknowledgement, trigger "DB302_HMI_Faults_Carrier59_Faults_0" bit 6
   3784: 'Carrier 59 PLC Not Communicating', class No Acknowledgement, trigger "DB302_HMI_Faults_Carrier59_Faults_0" bit 7
   3785: 'Carrier 59 Safe Input Card Fault', class No Acknowledgement, trigger "DB302_HMI_Faults_Carrier59_Faults_0" bit 8
   3786: 'Carrier 59 Safe Output Card Fault', class No Acknowledgement, trigger "DB302_HMI_Faults_Carrier59_Faults_0" bit 9
   3787: 'Carrier 59 Standard Input Card Fault', class No Acknowledgement, trigger "DB302_HMI_Faults_Carrier59_Faults_0" bit 10
   3788: 'Carrier 59 Standard Output Card Fault', class No Acknowledgement, trigger "DB302_HMI_Faults_Carrier59_Faults_0" bit 11
   3789: 'Carrier 59 Encoder Position Fault', class No Acknowledgement, trigger "DB302_HMI_Faults_Carrier59_Faults_0" bit 12
   3790: 'Carrier 59 Encoder Internal Error', class No Acknowledgement, trigger "DB302_HMI_Faults_Carrier59_Faults_0" bit 13
   3791: 'Carrier 59 Encoder Comm Fault', class No Acknowledgement, trigger "DB302_HMI_Faults_Carrier59_Faults_0" bit 14
   3792: 'Carrier 59 HMI Comm Fault', class No Acknowledgement, trigger "DB302_HMI_Faults_Carrier59_Faults_0" bit 15
   3793: 'Carrier 59 Crash Detection Fault', class No Acknowledgement, trigger "DB302_HMI_Faults_Carrier59_Faults_1" bit 0
   3794: 'Carrier 59 Carrier Number Invalid', class No Acknowledgement, trigger "DB302_HMI_Faults_Carrier59_Faults_1" bit 1
   3795: 'Carrier 59 Drive: PROFINET configuration error', class No Acknowledgement, trigger "DB302_HMI_Faults_Carrier59_Faults_1" bit 2
   3796: 'Carrier 59 Drive: Error internal communications', class No Acknowledgement, trigger "DB302_HMI_Faults_Carrier59_Faults_1" bit 3
   3797: 'Carrier 59 Drive: Motor overtemperature', class No Acknowledgement, trigger "DB302_HMI_Faults_Carrier59_Faults_1" bit 4
   3798: 'Carrier 59 Drive: Motor overcurrent', class No Acknowledgement, trigger "DB302_HMI_Faults_Carrier59_Faults_1" bit 5
   3799: 'Carrier 59 Drive: Infeed or power unit not ready', class No Acknowledgement, trigger "DB302_HMI_Faults_Carrier59_Faults_1" bit 6
   3800: 'Carrier 59 Drive: Short-circuit/ground fault detected', class No Acknowledgement, trigger "DB302_HMI_Faults_Carrier59_Faults_1" bit 7
   3801: 'Carrier 59 Drive: PROFINET Setpoint timeout', class No Acknowledgement, trigger "DB302_HMI_Faults_Carrier59_Faults_1" bit 8
   3802: 'Carrier 59 Power unit: Overcurrent', class No Acknowledgement, trigger "DB302_HMI_Faults_Carrier59_Faults_1" bit 9
   3803: 'Carrier 59 Power unit: DC link voltage overvoltage', class No Acknowledgement, trigger "DB302_HMI_Faults_Carrier59_Faults_1" bit 10
   3804: 'Carrier 59 Power unit: DC link voltage undervoltage', class No Acknowledgement, trigger "DB302_HMI_Faults_Carrier59_Faults_1" bit 11
   3805: 'Carrier 59 Power unit: Line phase failure in main circuit', class No Acknowledgement, trigger "DB302_HMI_Faults_Carrier59_Faults_1" bit 12
   3806: 'Carrier 59 Power unit: Phase failure motor cable', class No Acknowledgement, trigger "DB302_HMI_Faults_Carrier59_Faults_1" bit 13
   3807: 'Carrier 59 Power unit: Ground fault', class No Acknowledgement, trigger "DB302_HMI_Faults_Carrier59_Faults_1" bit 14
   3808: 'Spare_Fault_3808', class No Acknowledgement, trigger "DB302_HMI_Faults_Carrier59_Faults_1" bit 15
   3809: 'Carrier 59 Motion Off Fault', class No Acknowledgement, trigger "DB302_HMI_Faults_Carrier59_Faults_2" bit 0
   3810: 'Carrier 59 Motion On Fault', class No Acknowledgement, trigger "DB302_HMI_Faults_Carrier59_Faults_2" bit 1
   3811: 'Carrier 59 Spacing Fault', class No Acknowledgement, trigger "DB302_HMI_Faults_Carrier59_Faults_2" bit 2
   3812: 'Carrier 59 Duplicate Carrier Number Fault', class No Acknowledgement, trigger "DB302_HMI_Faults_Carrier59_Faults_2" bit 3
   3813: 'Spare_Fault_3813', class No Acknowledgement, trigger "DB302_HMI_Faults_Carrier59_Faults_2" bit 4
   3814: 'Spare_Fault_3814', class No Acknowledgement, trigger "DB302_HMI_Faults_Carrier59_Faults_2" bit 5